
     ELSIF (#tempPostfixNotation[#tempPositionOfPostfix] = #LGCODE_MTH_PRSR_LOGICAL_NOT) THEN
       IF #tempStackOfIntermediateResults[#tempPositionOfIntermediateResult - 1] <> 0 THEN
         #tempStackOfIntermediateResults[#tempPositionOfIntermediateResult - 1] := 0;
       ELSE
         #tempStackOfIntermediateResults[#tempPositionOfIntermediateResult - 1] := 1;
       END_IF;

     ELSIF (#tempPostfixNotation[#tempPositionOfPostfix] = #LGCODE_MTH_PRSR_LOGICAL_NOT_EQUAL) THEN
       IF
         #tempStackOfIntermediateResults[#tempPositionOfIntermediateResult - 2] <>
         #tempStackOfIntermediateResults[#tempPositionOfIntermediateResult - 1]
       THEN
         #tempStackOfIntermediateResults[#tempPositionOfIntermediateResult - 2] := 1;
       ELSE
         #tempStackOfIntermediateResults[#tempPositionOfIntermediateResult - 2] := 0;
       END_IF;
       #tempPositionOfIntermediateResult := #tempPositionOfIntermediateResult - 1;

     ELSIF (#tempPostfixNotation[#tempPositionOfPostfix] = #LGCODE_MTH_PRSR_LOGICAL_EQUAL) THEN
       IF
         #tempStackOfIntermediateResults[#tempPositionOfIntermediateResult - 2] =
         #tempStackOfIntermediateResults[#tempPositionOfIntermediateResult - 1]
       THEN
         #tempStackOfIntermediateResults[#tempPositionOfIntermediateResult - 2] := 1;
       ELSE
         #tempStackOfIntermediateResults[#tempPositionOfIntermediateResult - 2] := 0;
       END_IF;
       #tempPositionOfIntermediateResult := #tempPositionOfIntermediateResult - 1;

     ELSIF (#tempPostfixNotation[#tempPositionOfPostfix] = #LGCODE_MTH_PRSR_LOGICAL_AND) THEN
       IF
         #tempStackOfIntermediateResults[#tempPositionOfIntermediateResult - 2] > 0
         AND
         #tempStackOfIntermediateResults[#tempPositionOfIntermediateResult - 1] > 0
       THEN
         #tempStackOfIntermediateResults[#tempPositionOfIntermediateResult - 2] := 1;
       ELSE
         #tempStackOfIntermediateResults[#tempPositionOfIntermediateResult - 2] := 0;
       END_IF;
       #tempPositionOfIntermediateResult := #tempPositionOfIntermediateResult - 1;

     ELSIF (#tempPostfixNotation[#tempPositionOfPostfix] = #LGCODE_MTH_PRSR_LOGICAL_OR) THEN
       IF
         #tempStackOfIntermediateResults[#tempPositionOfIntermediateResult - 2] > 0
         OR
         #tempStackOfIntermediateResults[#tempPositionOfIntermediateResult - 1] > 0
       THEN
         #tempStackOfIntermediateResults[#tempPositionOfIntermediateResult - 2] := 1;
       ELSE
         #tempStackOfIntermediateResults[#tempPositionOfIntermediateResult - 2] := 0;
       END_IF;
       #tempPositionOfIntermediateResult := #tempPositionOfIntermediateResult - 1;

     END_IF;

     #tempPositionOfPostfix := #tempPositionOfPostfix + 1;

     #LKinLang_CalcMathAndBool.errorID := #LGCODE_MTH_PRSR_NO_ERR;
     #LKinLang_CalcMathAndBool.finalResult := #tempStackOfIntermediateResults[2];

   END_WHILE;

   //--------------------------------------------------------------------
   // End of Block LKinLang_CalcMathAndBool
   //--------------------------------------------------------------------
END_FUNCTION

FUNCTION "LKinLang_CharacterIsLetter" : Bool   // FC35454, SCL
TITLE = LKinLang_CharacterIsLetter
{ S7_Optimized_Access := 'TRUE' }
AUTHOR : tech.team.motioncontrol@siemens.com
FAMILY : LKinLang
VERSION : 1.1
// The FC checks a given character to be a letter
   VAR_INPUT
      character : Byte;   // character to be checked / character to be checked to be a letter
   END_VAR
   // Ret_Val : TRUE: character is letter; FALSE: character is NOT a letter
BEGIN
   //==========================================================================================
   // SIEMENS AG
   // (c)Copyright 2019 All Rights Reserved
   //------------------------------------------------------------------------------------------
   // Library: LKinLang
   // Tested with: S7-1517T-3 PN/DP
   // Engineering: TIA Portal V15
   // Restrictions: ---
   // Requirements: S7-1500T FW 2.5
   // Functionality: LKinLang_CharacterIsLetter
   // The FC checks a given character to be a letter 
   // 
   // Support: tech.team.motioncontrol@siemens.com
   // Note: Parameter comments are only available in language 'English (United States)'
   //------------------------------------------------------------------------------------------
   // Change log table:
   // Version    Date          Expert in charge    Changes applied
   // 01.00.00   28.05.2019    FR                  First created version
   // 01.01.00   09.01.2020    FR                  Added % as letter for interface vars
   //===========================================================================================

   //======================================================================
   // Check if the given characteracter is a LETTER
   //====================================================================== 

                      // A ..................... Z         
   IF ((#character >= 16#41 AND #character <= 16#5A) OR
                    // a ..................... z         
     (#character >= 16#61 AND #character <= 16#7A))
     OR #character = 16#25 //%
   THEN
     #LKinLang_CharacterIsLetter:= TRUE;
   ELSE
     #LKinLang_CharacterIsLetter := FALSE;
   END_IF;
END_FUNCTION

FUNCTION "LKinLang_CharacterIsMerger" : Bool   // FC35455, SCL
TITLE = LKinLang_CharacterIsMerger
{ S7_Optimized_Access := 'TRUE' }
AUTHOR : tech.team.motioncontrol@siemens.com
FAMILY : LKinLang
VERSION : 1.1
// The FC checks a given character to be a merger
   VAR_INPUT
      character : Byte;   // character to be checked
      lastIndexOfMerger : Int;
   END_VAR
   VAR_IN_OUT
      mergers : Array[1.."LKINLANG_NUMBER_OF_MERGERS"] of Byte;
   END_VAR
   VAR_TEMP
      tempCounter : Int;
   END_VAR
   // Ret_Val : TRUE: character is merger; FALSE: character is NOT a merger
BEGIN
   //==========================================================================================
   // SIEMENS AG
   // (c)Copyright 2019 All Rights Reserved
   //------------------------------------------------------------------------------------------
   // Library: LKinLang
   // Tested with: S7-1517T-3 PN/DP
   // Engineering: TIA Portal V15
   // Restrictions: ---
   // Requirements: S7-1500T FW 2.5
   // Functionality: LKinLang_CharacterIsMerger
   // The FC checks a given character to be a merger 
   // 
   // Support: tech.team.motioncontrol@siemens.com
   // Note: Parameter comments are only available in language 'English (United States)'
   //------------------------------------------------------------------------------------------
   // Change log table:
   // Version    Date          Expert in charge    Changes applied
   // 01.00.00   28.05.2019    FR                  First created version
   //===========================================================================================

   //======================================================================
   // Check if the given character is a merger
   //====================================================================== 

   #LKinLang_CharacterIsMerger := false;

   FOR #tempCounter := 1 TO #lastIndexOfMerger DO
     IF #mergers[#tempCounter] = #character THEN
       #LKinLang_CharacterIsMerger := true;
       EXIT;
     END_IF;
   END_FOR;
END_FUNCTION

FUNCTION "LKinLang_CharacterIsNumeric" : Bool   // FC35456, SCL
TITLE = LKinLang_CharacterIsNumeric
{ S7_Optimized_Access := 'TRUE' }
AUTHOR : tech.team.motioncontrol@siemens.com
FAMILY : LKinLang
VERSION : 1.1
// The FC checks a given character to be a numeric
   VAR_INPUT
      character : Char;   // character to be checked
   END_VAR
   // Ret_Val : TRUE: character is numeric; FALSE: character is NOT a numeric
BEGIN
   //==========================================================================================
   // SIEMENS AG
   // (c)Copyright 2019 All Rights Reserved
   //------------------------------------------------------------------------------------------
   // Library: LKinLang
   // Tested with: S7-1517T-3 PN/DP
   // Engineering: TIA Portal V15
   // Restrictions: ---
   // Requirements: S7-1500T FW 2.5
   // Functionality: LKinLang_CharacterIsNumeric
   // The FC checks a given character to be a numeric
   // 
   // Support: tech.team.motioncontrol@siemens.com
   // Note: Parameter comments are only available in language 'English (United States)'
   //------------------------------------------------------------------------------------------
   // Change log table:
   // Version    Date          Expert in charge    Changes applied
   // 01.00.00   28.05.2019    FR                  First created version
   //===========================================================================================

   //======================================================================
   // Check if the given character is a DIGIT or a POINT (used for comma)
   //====================================================================== 

   IF #character = '0'//16#30   // 0
     OR #character = '1'//16#31 // 1
     OR #character = '2'//16#32 // 2
     OR #character = '3'//16#33 // 3
     OR #character = '4'//16#34 // 4
     OR #character = '5'//16#35 // 5
     OR #character = '6'//16#36 // 6
     OR #character = '7'//16#37 // 7 
     OR #character = '8'//16#38 // 8
     OR #character = '9'//16#39 // 9 
     OR #character = '.'//16#2E // .
   THEN
     #LKinLang_CharacterIsNumeric := TRUE;
   ELSE
     #LKinLang_CharacterIsNumeric := FALSE;
   END_IF;
END_FUNCTION

FUNCTION "LKinLang_CheckLimits" : DWord   // FC35457, SCL
TITLE = LKinLang_CheckLimits
{ S7_Optimized_Access := 'TRUE' }
AUTHOR : tech.team.motioncontrol@siemens.com
FAMILY : LKinLang
VERSION : 1.1
// The FC checks a parameter value not to exceed give limits
   VAR_INPUT
      parameterMinVal : LReal;   // lower limit for parameter value
      parameterMaxVal : LReal;   // upper limit for parameter value
   END_VAR
   VAR_IN_OUT
      parameterValue : "LKinLang_typeDiffElementaryDatatypes";   // parameter value which is checked and written
   END_VAR
   VAR CONSTANT
      REAL_MIN : LReal := -3.402823E+38;
      REAL_MAX : LReal := 3.402823E+38;
      DINT_MIN : DInt := -2147483648;
      DINT_MAX : DInt := +2147483647;
      INT_MIN : Int := -32768;
      INT_MAX : Int := 32767;
      ERR_PARAMETER_OVERFLOW : DWord := 16#8000;
      ERR_PARAMETER_OUTSIDE_LIMITS : DWord := 16#8001;
   END_VAR
BEGIN
   //==========================================================================================
   // SIEMENS AG
   // (c)Copyright 2019 All Rights Reserved
   //------------------------------------------------------------------------------------------
   // Library: LKinLang
   // Tested with: S7-1517T-3 PN/DP
   // Engineering: TIA Portal V15
   // Restrictions: ---
   // Requirements: S7-1500T FW 2.5
   // Functionality: LKinLang_CheckLimits
   // The FC checks a parameter value not to exceed give limits
   // 
   // Support: tech.team.motioncontrol@siemens.com
   // Note: Parameter comments are only available in language 'English (United States)'
   //------------------------------------------------------------------------------------------
   // Change log table:
   // Version    Date          Expert in charge    Changes applied
   // 01.00.00   28.05.2019    FR                  First created version
   //===========================================================================================

   // ============================================================
   // Check limits of given parameter
   // ============================================================
   #LKinLang_CheckLimits := 0;

   // Check if parameter value is inside configured limits
   IF #parameterValue.valueLReal >= #parameterMinVal
     AND #parameterValue.valueLReal <= #parameterMaxVal
   THEN
     ; // Value is ok
   ELSE
     ; // Error: Value outside limits  
     #LKinLang_CheckLimits := #ERR_PARAMETER_OUTSIDE_LIMITS;
     RETURN;
   END_IF;

   // Check if parameter value (LReal) fits into smaller data types
   IF #parameterMinVal >= #REAL_MIN
     AND #parameterMaxVal <= #REAL_MAX
   THEN
     // Limits are OK
     IF #parameterValue.valueLReal <= #REAL_MAX
       AND #parameterValue.valueLReal >= #REAL_MIN
     THEN
       #parameterValue.valueReal := LREAL_TO_REAL(#parameterValue.valueLReal);
     ELSE
       // Error
       #LKinLang_CheckLimits := #ERR_PARAMETER_OVERFLOW;
       RETURN;
     END_IF;
   ELSE
     ;// Do nothing: because of the limits this format is not needed
   END_IF;

   IF #parameterMinVal >= #DINT_MIN
     AND #parameterMaxVal <= #DINT_MAX
   THEN
     // Limits are OK
     IF #parameterValue.valueLReal <= #DINT_MAX
       AND #parameterValue.valueLReal >= #DINT_MIN
     THEN
       #parameterValue.valueDint := LREAL_TO_DINT(#parameterValue.valueLReal);
     ELSE
       // Error
       #LKinLang_CheckLimits := #ERR_PARAMETER_OVERFLOW;
       RETURN;
     END_IF;
   ELSE
     ;// Do nothing: because of the limits this format is not needed
   END_IF;

   IF #parameterMinVal >= #INT_MIN
     AND #parameterMaxVal <= #INT_MAX
   THEN
     // Limits are OK
     IF #parameterValue.valueLReal <= #INT_MAX
       AND #parameterValue.valueLReal >= #INT_MIN
     THEN
       #parameterValue.valueInt := LREAL_TO_INT(#parameterValue.valueLReal);
     ELSE
       // Error
       #LKinLang_CheckLimits := #ERR_PARAMETER_OVERFLOW;
       RETURN;
     END_IF;
   ELSE
     ;// Do nothing: because of the limits this format is not needed
   END_IF;
END_FUNCTION

FUNCTION "LKinLang_CheckParameterCondition" : Bool   // FC35458, SCL
TITLE = LKinLang_CheckParameterCondition
{ S7_Optimized_Access := 'TRUE' }
AUTHOR : tech.team.motioncontrol@siemens.com
FAMILY : LKinLang
VERSION : 1.1
// The FC checks for conditions to be fullfilled
   VAR_INPUT
      mode : DInt;   // Selected mode, where the parameters are to be checked (0: In line, 1: In Cmd, 2: In Prg)
      language : Int;   // Selected language
   END_VAR
   VAR_OUTPUT
      errorString : String;   // Generated error message
   END_VAR
   VAR_IN_OUT
      setParameters : Array[1.."LKINLANG_NUMBER_OF_CONDITIONS"] of "LKinLang_typeCondition";   // Array containint all parameters which are set for the selected mode
      conditionsToCheck : Array[1.."LKINLANG_NUMBER_OF_CONDITIONS"] of "LKinLang_typeCondition";   // Array containing all parameters which are to be checked
      parameterDefaults : Variant;   // Parameter defaults to call SelectLangPackage
   END_VAR
   VAR_TEMP
      tempParameterOk : Bool;   // Temporary variable for the return value of this FC
      tempGroupToCheck : DInt;   // Temporary variable for the group which is checked
      tempParameterToCheck : DInt;   // Temporary variable for the parameter number which is checked
      tempConditionCounter : Int;   // Temporary counter in the conditions array
      tempSetCounter : Int;   // Temporary counter in the parameters array
      tempConditionUpperLimit : DInt;   // Temporary variable for upper limit of conditions array
      tempConditionLowerLimit : DInt;   // Temporary variable for lower limit of conditions array
      tempSetUpperLimit : DInt;   // Temporary variable for upper limit of parameters array
      tempSetLowerLimit : DInt;   // Temporary variable for lower limit of parameters array
      tempGroups : Array[1.."LKINLANG_NUMBER_OF_CONDITIONS"] of DInt;   // Temporay array for all groups to be checked
      tempGroupCounter : DInt;   // Temporary variable for last entry in groups array
      tempCounter : Int;   // Temporary counter
      tempParameterDefinition : "LKinLang_typeParameterDefinition";   // Temporary variable for the parameter definition
      tempSep : Array[1.."LKINLANG_NUMBER_OF_SEPARATORS"] of Byte;   // Temporary variable for separators array
      tempMerg : Array[1.."LKINLANG_NUMBER_OF_MERGERS"] of Byte;   // Temporary variable for mergers array
      tempValidCounts : "LKinLang_typePathDataElementCounter";   // Temporary variable for valid counts array
      tempString : "LKinLang_typeVariableDeclaration";
      tempKeyToken : "LKinLang_typeKeyToken";
   END_VAR
   // Ret_Val : Return value of this FC
BEGIN
   //==========================================================================================
   // SIEMENS AG
   // (c)Copyright 2019 All Rights Reserved
   //------------------------------------------------------------------------------------------
   // Library: LKinLang
   // Tested with: S7-1517T-3 PN/DP
   // Engineering: TIA Portal V15
   // Restrictions: ---
   // Requirements: S7-1500T FW 2.5
   // Functionality: LKinLang_CheckParameterCondition
   // This function searches the array "SetParameters" if the parameter number from "ConditionsToCheck" is set.
   // For each group ("conditionsToCheck.Group") there must be at least one parameter number in "SetParameters".
   // 
   // The mode to check is given as an Input:
   // 0: "SetParameters" in the actual line are checked
   // 1: "SetParameters" in the actual command are checked
   // 2: "SetParameters" in the complete program are checked
   // The respective "SetParameters" array must be connected outside
   // 
   // Support: tech.team.motioncontrol@siemens.com
   // Note: Parameter comments are only available in language 'English (United States)'
   //------------------------------------------------------------------------------------------
   // Change log table:
   // Version    Date          Expert in charge    Changes applied
   // 01.00.00   28.05.2019    FR                  First created version
   //===========================================================================================

   // Init variables
   #tempParameterOk := #LKinLang_CheckParameterCondition := FALSE;
   #tempGroupCounter := 0;

   // Get limits of "conditionToCheck" array
   #tempConditionLowerLimit := 1;
   #tempConditionUpperLimit := "LKINLANG_NUMBER_OF_CONDITIONS";

   // Get limits of "setParameters" array
   #tempSetLowerLimit := 1;
   #tempSetUpperLimit := "LKINLANG_NUMBER_OF_CONDITIONS";

   // Iterate over condition array and get all groups which are to be checked
   FOR #tempCounter := #tempConditionLowerLimit TO #tempConditionUpperLimit DO
     // Get group to check
     IF #conditionsToCheck[#tempCounter].Group <> 0 // Group is not 0
       AND #tempGroupToCheck <> #conditionsToCheck[#tempCounter].Group // Group is different from already added group
       AND #conditionsToCheck[#tempCounter].Mode = #mode // Mode is same as selected input
     THEN
       // Increment counter for found groups 
       #tempGroupCounter += 1;
       // Save group number in temp for check in next iteration
       #tempGroupToCheck := #conditionsToCheck[#tempCounter].Group;
       // Save group in array to work with later
       #tempGroups[#tempGroupCounter] := #conditionsToCheck[#tempCounter].Group;
     END_IF;
   END_FOR;

   // Iterate over all found groups ("tempGroups")
   FOR #tempCounter := 1 TO #tempGroupCounter DO
     // Reset Parameter ok
     #tempParameterOk := FALSE;
     // Reset parameter number to check
     #tempParameterToCheck := -1;

     // Search if one group member (parameterNumber) is in "SetParameters" Array 
     FOR #tempConditionCounter := #tempConditionLowerLimit TO #tempConditionUpperLimit DO

       // Search for entries in conditionsToCheck array where ".Group" fits "tempGroups" 
       IF #conditionsToCheck[#tempConditionCounter].Group = #tempGroups[#tempCounter] THEN
         // Group is same --> Get parameter number to check
         #tempParameterToCheck := #conditionsToCheck[#tempConditionCounter].ParameterNumber;
       END_IF;

       // Search in array "SetParameters" if there is an entry which fits the parameterToCheck
       FOR #tempSetCounter := #tempSetLowerLimit TO #tempSetUpperLimit DO
         IF #tempParameterToCheck = #setParameters[#tempSetCounter].ParameterNumber THEN
           // Parameter number was found --> Set parameter ok to True and exit this for Loop
           #tempParameterOk := true;
           EXIT;
         END_IF;
       END_FOR;

       // If one of the group members was found also exit this for loop
       IF #tempParameterOk THEN
         EXIT;
       END_IF;
     END_FOR;

     // If parameter number was not found, generate error message
     IF NOT #tempParameterOk THEN
       // Parameter / Group is missing 
       #errorString := 'Mandatory parameter ';

       FOR #tempConditionCounter := #tempConditionLowerLimit TO #tempConditionUpperLimit DO
         // Get parameter number in conditions to check array, where group fits
         IF #conditionsToCheck[#tempConditionCounter].Group = #tempGroups[#tempCounter] THEN

           // Copy found parameter number
           #tempParameterToCheck := #conditionsToCheck[#tempConditionCounter].ParameterNumber;

           // Get definition of parameter with this number
           "LKinLang_SelectLangPackage"(language := #language,
                                        variableDeclarations=>#tempString,
                                        keyToken=>#tempKeyToken,
                                        parameterDefinition := #tempParameterDefinition,
                                        separators => #tempSep,
                                        mergers => #tempMerg,
                                        validCounts => #tempValidCounts,
                                        parameterNumber := #tempParameterToCheck,
                                        parameterDefaults := #parameterDefaults);


           // Copy the name of the parameter to the error string
           #errorString := CONCAT(IN1 := #errorString, IN2 := #tempParameterDefinition.parameterNameString);

           IF #tempParameterDefinition.parameterNameNumber <> -1 THEN
             // Concat parameterNameNumber and delete sign from DINT_TO_STRING
             #errorString := CONCAT(IN1 := #errorString, IN2 := DELETE(IN := DINT_TO_STRING(#tempParameterDefinition.parameterNameNumber), L := 1, P := 1));
           END_IF;
           // Seperate parameters from the same group with ", "
           #errorString := CONCAT(IN1 := #errorString, IN2 := ', ');
         END_IF;

       END_FOR;
       // Delete last ", "
       #errorString := LEFT(IN := #errorString, L := LEN(#errorString) - 2);
       // Concat last strings
       #errorString := CONCAT(IN1 := #errorString, IN2 := ' is missing');
       // The resulting errorString should look like this
       // "Mandatory parameter G17, G18, G19 is missing" (G17, G18, G19 are for example in the same condition group)
       // 
       // Return from this function
       RETURN;

     ELSE
       // Reset parameter ok for the next group to check
       #tempParameterOk := false;
     END_IF;

   END_FOR;

   // If all groups are ok set parameterOk to true
   // We can assume all parameters were ok because else we would have returned after writing the error string
   #tempParameterOk := true;

   // Write internal temp to output
   #LKinLang_CheckParameterCondition := #tempParameterOk;

   //===========================================================================================
   // End of Block
   //===========================================================================================
END_FUNCTION

FUNCTION "LKinLang_CheckParameterCounter" : Void   // FC35459, SCL
TITLE = LKinLang_CheckParameterCounter
{ S7_Optimized_Access := 'TRUE' }
AUTHOR : tech.team.motioncontrol@siemens.com
FAMILY : LKinLang
VERSION : 1.1
// This function checks how often a parameter was programmed in one line
   VAR_INPUT
      parameterNumber : Int;   // Parameter number for which the counter is checked
      lineNo : UInt;   // Actual line number for error message
      parameterDefinition : "LKinLang_typeParameterDefinition";   // Parameter definition of the parameter number
   END_VAR
   VAR_IN_OUT
      parameterCounter : Array[*] of "LKinLang_typeParameterCounter";   // Parameter counter array
      errorString : String;   // Error message
      error : Bool;   // Error output
   END_VAR
   VAR_TEMP
      tempCounter : Int;   // Temporary counter
      tempUBound : DInt;   // Temporary variable for the upper limit of the parameterCounter array
      tempLBound : DInt;   // Temporary variable for the lower limit of the parameterCounter array
      tempParameterFound : Bool;   // Temporary bit to signalize if the parameter is already in the parameterCounter array
   END_VAR
   // Ret_Val : No return value
BEGIN
   //==========================================================================================
   // SIEMENS AG
   // (c)Copyright 2019 All Rights Reserved
   //------------------------------------------------------------------------------------------
   // Library: LKinLang
   // Tested with: S7-1517T-3 PN/DP
   // Engineering: TIA Portal V15
   // Restrictions: ---
   // Requirements: S7-1500T FW 2.5
   // Functionality: LKinLang_CheckParameterCounter
   // This function checks how often a given parameter was programmed in one line.
   // It increases the counter or throws an error if the limit is exceeded.
   //
   // Support: tech.team.motioncontrol@siemens.com
   // Note: Parameter comments are only available in language 'English (United States)'
   //------------------------------------------------------------------------------------------
   // Change log table:
   // Version    Date          Expert in charge    Changes applied
   // 01.00.00   28.05.2019    FR                  First created version
   //===========================================================================================

   // Initialize variables
   //------------------------------------------------------------------------------------------
   #tempLBound := LOWER_BOUND(ARR := #parameterCounter, DIM := 1);
   #tempUBound := UPPER_BOUND(ARR := #parameterCounter, DIM := 1);
   #tempParameterFound := FALSE;
   //------------------------------------------------------------------------------------------

   // Check if parameter number is already in array
   //------------------------------------------------------------------------------------------
   FOR #tempCounter := #tempLBound TO #tempUBound DO

     // Parameter number is already in array
     IF #parameterCounter[#tempCounter].parameterNumber = #parameterNumber THEN

       // Already in array --> Count up
       #parameterCounter[#tempCounter].counterValue += 1;
       // Set bit to skip creating a new entry
       #tempParameterFound := TRUE;

       // ERROR: Throw error if limit of counter was exceeded
       //------------------------------------------------------------------------------------------
       IF #parameterCounter[#tempCounter].counterValue > #parameterDefinition.validCountPerLine THEN

         // Create error string
         //------------------------------------------------------------------------------------------
         #errorString := CONCAT(IN1 := #errorString, IN2 := 'Programmed ');
         #errorString := CONCAT(IN1 := #errorString, IN2 := #parameterDefinition.parameterNameString);

         // Concat parameterNameNumber if not -1
         // If the parameter does not include a number, e.g. LIN (compared to G2) the parameterNameNumber is -1 by default 
         IF #parameterDefinition.parameterNameNumber <> -1 THEN
           #errorString := CONCAT(IN1 := #errorString, IN2 := DINT_TO_STRING(#parameterDefinition.parameterNameNumber));
         END_IF;
         #errorString := CONCAT(IN1 := #errorString, IN2 := ' too often: Allowed:');
         #errorString := CONCAT(IN1 := #errorString, IN2 := DINT_TO_STRING(#parameterDefinition.validCountPerLine));
         #errorString := CONCAT(IN1 := #errorString, IN2 := ' Programmed:');
         #errorString := CONCAT(IN1 := #errorString, IN2 := INT_TO_STRING(#parameterCounter[#tempCounter].counterValue));
         #errorString := CONCAT(IN1 := #errorString, IN2 := '; Line:');
         #errorString := CONCAT(IN1 := #errorString, IN2 := UINT_TO_STRING(#lineNo));

         // Completed errorString should look like
         // "Programmed G1 too often: Allowed:+1 Programmed: +2; Line:+10 "
         //------------------------------------------------------------------------------------------

         // Set error output to TRUE;
         #error := TRUE;

         // Return from function after errorString is written
         RETURN;
       ELSE
         // Exit for loop if parameter was found and counter was sucessfully increased
         EXIT;
       END_IF;
     ELSE
       ; // Do nothing --> next iteration
     END_IF;
   END_FOR;
   //------------------------------------------------------------------------------------------

   // If parameter was not found, create new entry in parameterCounter array
   //------------------------------------------------------------------------------------------
   IF NOT #tempParameterFound THEN
     // New entry
     // Search empty array index
     FOR #tempCounter := #tempLBound TO #tempUBound DO

       // If CounterValue = 0 then this must be a empty index
       IF #parameterCounter[#tempCounter].counterValue = 0 THEN

         // New entry
         #parameterCounter[#tempCounter].parameterNumber := #parameterNumber;
         // Increment counter
         #parameterCounter[#tempCounter].counterValue += 1;

         // ERROR: Throw error if limit of counter was exceeded
         //------------------------------------------------------------------------------------------
         IF #parameterCounter[#tempCounter].counterValue > #parameterDefinition.validCountPerLine THEN

           // Create error string
           //------------------------------------------------------------------------------------------
           #errorString := CONCAT(IN1 := #errorString, IN2 := 'Programmed ');
           #errorString := CONCAT(IN1 := #errorString, IN2 := #parameterDefinition.parameterNameString);
           // Concat parameterNameNumber if not -1
           // If the parameter does not include a number, e.g. LIN (compared to G2) the parameterNameNumber is -1 by default 
           IF #parameterDefinition.parameterNameNumber <> -1 THEN
             #errorString := CONCAT(IN1 := #errorString, IN2 := DINT_TO_STRING(#parameterDefinition.parameterNameNumber));
           END_IF;
           #errorString := CONCAT(IN1 := #errorString, IN2 := ' too often: Allowed:');
           #errorString := CONCAT(IN1 := #errorString, IN2 := DINT_TO_STRING(#parameterDefinition.validCountPerLine));
           #errorString := CONCAT(IN1 := #errorString, IN2 := ' Programmed:');
           #errorString := CONCAT(IN1 := #errorString, IN2 := INT_TO_STRING(#parameterCounter[#tempCounter].counterValue));
           #errorString := CONCAT(IN1 := #errorString, IN2 := '; Line:');
           #errorString := CONCAT(IN1 := #errorString, IN2 := UINT_TO_STRING(#lineNo));

           // Completed errorString should look like
           // "Programmed G1 too often: Allowed:+1 Programmed: +2; Line:+10 "
           //------------------------------------------------------------------------------------------

           // Set error output to TRUE;
           #error := TRUE;

           // Return from function after errorString is written
           RETURN;
         ELSE
           // Exit for loop if parameter was found and counter was sucessfully increased
           EXIT;
         END_IF;
       ELSE
         ; // Do nothing --> next iteration
       END_IF;
     END_FOR;
     //------------------------------------------------------------------------------------------
   ELSE
     ; // Do nothing --> parameter was found before
   END_IF;

   //===========================================================================================
   // End of Block
   //===========================================================================================
END_FUNCTION

FUNCTION "LKinLang_CheckPathDataCmd" : Word   // FC35460, SCL
TITLE = LKinCtrl_CheckPathDataCmd
{ S7_Optimized_Access := 'TRUE' }
AUTHOR : tech.team.motioncontrol@siemens.com
FAMILY : LKinCtrl
VERSION : 1.1
// The FC checks a PathData command to be configured correctly
   VAR_IN_OUT
      errorString : String;
      pathDataCmd : "LKinCtrl_typePathDataElement_advanced";   // variant for PathData command
   END_VAR
   VAR_TEMP
      tmpError : Bool;   // temporary variable for error bit
      tempFlagCtr : Int;   // temporary counter for flags
   END_VAR
   VAR CONSTANT
      STATUS_NO_ERROR_IN_COMMAND : Word := 16#0000;   // status no error found command
      ERR_PATHDATA_CMDTYPE : Word := 16#80A0;   // error due to wrong cmdType
      ERR_PATHDATA_COORDSYSTEM : Word := 16#80B1;   // error due to wrong coordinate system
      ERR_PATHDATA_ORIENTATIONDIRECTION : Word := 16#8007;   // error due to wrong orientation direction
      ERR_PATHDATA_BUFFERMODE : Word := 16#80B2;   // error due to wrong buffer mode
      ERR_PATHDATA_DYNAMICADAPTION : Word := 16#80B5;   // error due to wrong dynamic adaption
      ERR_PATHDATA_CIRCMODE : Word := 16#80B6;   // error due to wrong circle mode
      ERR_PATHDATA_PATHCHOICE : Word := 16#80B9;   // error due to wrong path choice
      ERR_PATHDATA_CIRCLEPLANE : Word := 16#80BA;   // error due to wrong circle plane
      ERR_PATHDATA_RADIUS : Word := 16#80BB;   // error due to wrong radius
      ERR_PATHDATA_ARC : Word := 16#80BC;   // error due to wrong arc
      ERR_PATHDATA_SETFLAGS_FLAG : Word := 16#80D1;   // error due to wrong flag definition
      ERR_PATHDATA_SETFLAGS_FLAGMODE : Word := 16#80D2;   // error due to wrong flag mode definition / errot due to wrong flag mode definition
      ERR_PATHDATA_OFFSET_PARA_NO : Word := 16#80A1;   // error due to wrong offset parameter set number / errot due to wrong offset parameter set number
      ERR_PATHDATA_OFFSET_MAINPATHPLANE : Word := 16#80A2;   // error due to wrong main path plane
      MINVAL_LREAL : LReal := -1.7976931348623157E+308;
      MINVAL_DINT : DInt := -2_147_483_648;
      MINVAL_INT : Int := -32_768;
   END_VAR
BEGIN
   //==========================================================================================
   // SIEMENS AG
   // (c)Copyright 2019 All Rights Reserved
   //------------------------------------------------------------------------------------------
   // Library: LKinLang
   // Tested with: S7-1517T-3 PN/DP
   // Engineering: TIA Portal V15
   // Restrictions: ---
   // Requirements: S7-1500T FW 2.5
   // Functionality: LKinLang_CheckPathDataCmd
   // The FC checks a PathData command to be configured correctly
   // 
   // Support: tech.team.motioncontrol@siemens.com
   // Note: Parameter comments are only available in language 'English (United States)'
   //------------------------------------------------------------------------------------------
   // Change log table:
   // Version    Date          Expert in charge    Changes applied
   // 01.00.00   28.05.2019    FR                  First created version
   // 01.00.01   26.11.2019    FR                  Added flagOnly cmd to CmdType check; added value Flags
   // 01.00.02   12.02.2020    FR                  Use correct constant for valueFlags
   // 01.00.03   10.12.2020    FR                  Check for cmdType=-1 
   //===========================================================================================

   // FC initialization
   //====================================================================================================================================
   #tmpError := FALSE;
   #LKinLang_CheckPathDataCmd := #STATUS_NO_ERROR_IN_COMMAND;

   // PathData command 
   //====================================================================================================================================
   //PathData - command - cmdType
   // Check for cmdType = -1 
   // This FC is only called to check valid motion commands
   // => -1 is not allowed
   // => End of PathData is written in other step
   IF #pathDataCmd.cmdType = -1 THEN
       #tmpError := TRUE;
       #LKinLang_CheckPathDataCmd := #ERR_PATHDATA_CMDTYPE;
       #errorString := CONCAT(IN1 := #errorString, IN2 := 'Error: Missing motion command');
       RETURN;
   END_IF;


   // check for wrong PathData parameter cmdType
   IF (#pathDataCmd.cmdType < "LKINCTRL_CMD_FLAG_ONLY"                      // lower limit MC cmdTypes
     OR #pathDataCmd.cmdType > "LKINCTRL_MC_MOVECIRCULARREL")               // upper limit MC cmdTypes
     AND #pathDataCmd.cmdType <> "LKINCTRL_CMD_WAIT_TIME"                   // exact cmdType constant for wait time
     AND #pathDataCmd.cmdType <> "LKINCTRL_CONFIG_START_OFFSET_COMP_LEFT"   // exact cmdType constant for activation offset compensation left
     AND #pathDataCmd.cmdType <> "LKINCTRL_CONFIG_START_OFFSET_COMP_RIGHT"  // exact cmdType constant for activation offset compensation right
     AND #pathDataCmd.cmdType <> "LKINCTRL_CONFIG_END_OFFSET_COMP"          // exact cmdType constant for deactivation offset compensation
   THEN
     #tmpError := TRUE;
     #LKinLang_CheckPathDataCmd := #ERR_PATHDATA_CMDTYPE;
     #errorString := CONCAT(IN1 := #errorString, IN2 := 'Error: cmdType = ');
     #errorString := CONCAT(IN1 := #errorString, IN2 := INT_TO_STRING(#pathDataCmd.cmdType));
     #errorString := CONCAT(IN1 := #errorString, IN2 := ' not allowed');
     RETURN;
   END_IF;


   //PathData - command - cmdCoordinates - coordSystem
   // check for wrong parameter PathData coordSystem
   IF #pathDataCmd.cmdCoordinates.coordSystem < 0
     AND #pathDataCmd.cmdCoordinates.coordSystem > 3
   THEN
     #tmpError := TRUE;
     #LKinLang_CheckPathDataCmd := #ERR_PATHDATA_COORDSYSTEM;
     #errorString := CONCAT(IN1 := #errorString, IN2 := 'Error: Coordinate system = ');
     #errorString := CONCAT(IN1 := #errorString, IN2 := DINT_TO_STRING(#pathDataCmd.cmdCoordinates.coordSystem));
     #errorString := CONCAT(IN1 := #errorString, IN2 := ' not allowed');
     RETURN;
   END_IF;

   //PathData - command - cmdParameters - orientationDirection
   // check for wrong parameter PathData orientationDirection
   IF #pathDataCmd.cmdParameters.orientationDirection < 1
     OR #pathDataCmd.cmdParameters.orientationDirection > 3
   THEN
     #tmpError := TRUE;
     #LKinLang_CheckPathDataCmd := #ERR_PATHDATA_ORIENTATIONDIRECTION;
     #errorString := CONCAT(IN1 := #errorString, IN2 := 'Error: Orientation direction = ');
     #errorString := CONCAT(IN1 := #errorString, IN2 := DINT_TO_STRING(#pathDataCmd.cmdParameters.orientationDirection));
     #errorString := CONCAT(IN1 := #errorString, IN2 := ' not allowed');
     RETURN;
   END_IF;

   //PathData - command - cmdParameters - bufferMode
   // check for wrong parameter PathData bufferMode
   IF #pathDataCmd.cmdParameters.bufferMode <> 1
     AND #pathDataCmd.cmdParameters.bufferMode <> 2
     AND #pathDataCmd.cmdParameters.bufferMode <> 5
   THEN
     #tmpError := TRUE;
     #LKinLang_CheckPathDataCmd := #ERR_PATHDATA_BUFFERMODE;
     #errorString := CONCAT(IN1 := #errorString, IN2 := 'Error: Buffer mode = ');
     #errorString := CONCAT(IN1 := #errorString, IN2 := DINT_TO_STRING(#pathDataCmd.cmdParameters.bufferMode));
     #errorString := CONCAT(IN1 := #errorString, IN2 := ' not allowed');
     RETURN;
   END_IF;

   //PathData - command - cmdParameters - dynamicAdaption
   // check for wrong parameter PathData dynamicAdaption
   IF #pathDataCmd.cmdParameters.dynamicAdaption > 2
   THEN
     #tmpError := TRUE;
     #LKinLang_CheckPathDataCmd := #ERR_PATHDATA_DYNAMICADAPTION;
     #errorString := CONCAT(IN1 := #errorString, IN2 := 'Error: Dynamic adaption = ');
     #errorString := CONCAT(IN1 := #errorString, IN2 := DINT_TO_STRING(#pathDataCmd.cmdParameters.dynamicAdaption));
     #errorString := CONCAT(IN1 := #errorString, IN2 := ' not allowed');
     RETURN;
   END_IF;

   //PathData - command - circleParameter
   //====================================================================================================================================
   //PathData - command - circleParameter - circMode
   // check for wrong parameter PathData circMode
   IF #pathDataCmd.cmdParameters.circleParameters.circMode < 0
     OR #pathDataCmd.cmdParameters.circleParameters.circMode > 3
   THEN
     #tmpError := TRUE;
     #LKinLang_CheckPathDataCmd := #ERR_PATHDATA_CIRCMODE;
     #errorString := CONCAT(IN1 := #errorString, IN2 := 'Error: Circle mode = ');
     #errorString := CONCAT(IN1 := #errorString, IN2 := DINT_TO_STRING(#pathDataCmd.cmdParameters.circleParameters.circMode));
     #errorString := CONCAT(IN1 := #errorString, IN2 := ' not allowed');
     RETURN;
   END_IF;

   //PathData - command - circleParameter - pathChoice
   // check for wrong parameter PathData pathChoice
   IF #pathDataCmd.cmdParameters.circleParameters.pathChoice < 0
     OR #pathDataCmd.cmdParameters.circleParameters.pathChoice > 3
   THEN
     #tmpError := TRUE;
     #LKinLang_CheckPathDataCmd := #ERR_PATHDATA_PATHCHOICE;
     #errorString := CONCAT(IN1 := #errorString, IN2 := 'Error: Path choice = ');
     #errorString := CONCAT(IN1 := #errorString, IN2 := DINT_TO_STRING(#pathDataCmd.cmdParameters.circleParameters.pathChoice));
     #errorString := CONCAT(IN1 := #errorString, IN2 := ' not allowed');
     RETURN;
   END_IF;

   //PathData - command - circleParameter - circlePlane
   // check for wrong parameter PathData circlePlane
   IF #pathDataCmd.cmdParameters.circleParameters.circlePlane < 0
     OR #pathDataCmd.cmdParameters.circleParameters.circlePlane > 2
   THEN
     #tmpError := TRUE;
     #LKinLang_CheckPathDataCmd := #ERR_PATHDATA_CIRCLEPLANE;
     #errorString := CONCAT(IN1 := #errorString, IN2 := 'Error: Circle plane = ');
     #errorString := CONCAT(IN1 := #errorString, IN2 := DINT_TO_STRING(#pathDataCmd.cmdParameters.circleParameters.circlePlane));
     #errorString := CONCAT(IN1 := #errorString, IN2 := ' not allowed');
     RETURN;
   END_IF;

   //PathData - command - circleParameter - radius
   // check for wrong parameter PathData radius
   IF #pathDataCmd.cmdParameters.circleParameters.radius < 0.0
   THEN
     #tmpError := TRUE;
     #LKinLang_CheckPathDataCmd := #ERR_PATHDATA_RADIUS;
     #errorString := CONCAT(IN1 := #errorString, IN2 := 'Error: Circle radius = ');
     #errorString := CONCAT(IN1 := #errorString, IN2 := LREAL_TO_STRING(#pathDataCmd.cmdParameters.circleParameters.radius));
     #errorString := CONCAT(IN1 := #errorString, IN2 := ' not allowed');
     RETURN;
   END_IF;

   //PathData - command - circleParameter - arc
   // check for wrong parameter PathData arc
   IF #pathDataCmd.cmdParameters.circleParameters.arc < 0.0
   THEN
     #tmpError := TRUE;
     #LKinLang_CheckPathDataCmd := #ERR_PATHDATA_ARC;
     #errorString := CONCAT(IN1 := #errorString, IN2 := 'Error: Circle arc = ');
     #errorString := CONCAT(IN1 := #errorString, IN2 := LREAL_TO_STRING(#pathDataCmd.cmdParameters.circleParameters.arc));
     #errorString := CONCAT(IN1 := #errorString, IN2 := ' not allowed');
     RETURN;
   END_IF;

   //PathData - command - offsetParameters - offSetParaNo
   // check for wrong parameter offSetParaNo
   IF (#pathDataCmd.cmdType = "LKINCTRL_CONFIG_START_OFFSET_COMP_LEFT"
     OR #pathDataCmd.cmdType = "LKINCTRL_CONFIG_START_OFFSET_COMP_RIGHT")
     AND (#pathDataCmd.cmdParameters.offsetParameters.offsetParaNo < 1
     OR #pathDataCmd.cmdParameters.offsetParameters.offsetParaNo > "LKINCTRL_NO_OF_OFFSETS")
   THEN
     #tmpError := TRUE;
     #LKinLang_CheckPathDataCmd := #ERR_PATHDATA_OFFSET_PARA_NO;
     #errorString := CONCAT(IN1 := #errorString, IN2 := 'Error: Offset parameter number = ');
     #errorString := CONCAT(IN1 := #errorString, IN2 := DINT_TO_STRING(#pathDataCmd.cmdParameters.offsetParameters.offsetParaNo));
     #errorString := CONCAT(IN1 := #errorString, IN2 := ' not allowed');
     RETURN;
   END_IF;

   //PathData - command - offsetParameters - main
   // check for wrong parameter PathData circlePlane
   IF (#pathDataCmd.cmdType = "LKINCTRL_CONFIG_START_OFFSET_COMP_LEFT"
     OR #pathDataCmd.cmdType = "LKINCTRL_CONFIG_START_OFFSET_COMP_RIGHT")
     AND (#pathDataCmd.cmdParameters.offsetParameters.mainPathPlane < 0
     OR #pathDataCmd.cmdParameters.offsetParameters.mainPathPlane > 2)
   THEN
     #tmpError := TRUE;
     #LKinLang_CheckPathDataCmd := #ERR_PATHDATA_OFFSET_MAINPATHPLANE;
     #errorString := CONCAT(IN1 := #errorString, IN2 := 'Error: Offset main path plane = ');
     #errorString := CONCAT(IN1 := #errorString, IN2 := DINT_TO_STRING(#pathDataCmd.cmdParameters.offsetParameters.mainPathPlane));
     #errorString := CONCAT(IN1 := #errorString, IN2 := ' not allowed');
     RETURN;
   END_IF;

   //PathData - command - setFlags
   //====================================================================================================================================
   FOR #tempFlagCtr := 1 TO "LKINCTRL_NO_OF_CMD_SETFLAGS" DO
     // check flag to be in range of flags InOut array at LKinCtrl_MC_MovePath
     IF #pathDataCmd.setFlags[#tempFlagCtr].flag < -1
       OR #pathDataCmd.setFlags[#tempFlagCtr].flag > "LKINCTRL_NO_OF_LAST_SETFLAG"
     THEN
       #tmpError := TRUE;
       #LKinLang_CheckPathDataCmd := #ERR_PATHDATA_SETFLAGS_FLAG;
       #errorString := CONCAT(IN1 := #errorString, IN2 := 'Error: Flag index = ');
       #errorString := CONCAT(IN1 := #errorString, IN2 := DINT_TO_STRING(#pathDataCmd.setFlags[#tempFlagCtr].flag));
       #errorString := CONCAT(IN1 := #errorString, IN2 := ' not allowed');
       EXIT;
       RETURN;
     END_IF;

     // check flagMode to be valid
     IF #pathDataCmd.setFlags[#tempFlagCtr].flagMode <> 0
       AND #pathDataCmd.setFlags[#tempFlagCtr].flagMode <> 1
       AND #pathDataCmd.setFlags[#tempFlagCtr].flagMode <> 2
       AND #pathDataCmd.setFlags[#tempFlagCtr].flagMode <> 3
       AND #pathDataCmd.setFlags[#tempFlagCtr].flagMode <> 5
       AND #pathDataCmd.setFlags[#tempFlagCtr].flagMode <> 10
       AND #pathDataCmd.setFlags[#tempFlagCtr].flagMode <> 11
       AND #pathDataCmd.setFlags[#tempFlagCtr].flagMode <> 13
       AND #pathDataCmd.setFlags[#tempFlagCtr].flagMode <> 15
     THEN
       #tmpError := TRUE;
       #LKinLang_CheckPathDataCmd := #ERR_PATHDATA_SETFLAGS_FLAGMODE;
       #errorString := CONCAT(IN1 := #errorString, IN2 := 'Error: Flag mode = ');
       #errorString := CONCAT(IN1 := #errorString, IN2 := DINT_TO_STRING(#pathDataCmd.setFlags[#tempFlagCtr].flagMode));
       #errorString := CONCAT(IN1 := #errorString, IN2 := ' not allowed');
       EXIT;
       RETURN;
     END_IF;
   END_FOR;

   //PathData - command - valueFlags
   //====================================================================================================================================
   FOR #tempFlagCtr := 1 TO "LKINCTRL_NO_OF_CMD_VALUEFLAGS" DO
     // check flag to be in range of flags InOut array at LKinCtrl_MC_MovePath
     IF #pathDataCmd.valueFlags[#tempFlagCtr].flag < -1
       OR #pathDataCmd.valueFlags[#tempFlagCtr].flag > "LKINCTRL_NO_OF_LAST_VALUEFLAG"
     THEN
       #tmpError := TRUE;
       #LKinLang_CheckPathDataCmd := #ERR_PATHDATA_SETFLAGS_FLAG;
       #errorString := CONCAT(IN1 := #errorString, IN2 := 'Error: Flag index = ');
       #errorString := CONCAT(IN1 := #errorString, IN2 := DINT_TO_STRING(#pathDataCmd.valueFlags[#tempFlagCtr].flag));
       #errorString := CONCAT(IN1 := #errorString, IN2 := ' not allowed');
       EXIT;
       RETURN;
     END_IF;

     // check flagMode to be valid
     IF #pathDataCmd.valueFlags[#tempFlagCtr].flagMode <> 0
       AND #pathDataCmd.valueFlags[#tempFlagCtr].flagMode <> 1
       AND #pathDataCmd.valueFlags[#tempFlagCtr].flagMode <> 2
       AND #pathDataCmd.valueFlags[#tempFlagCtr].flagMode <> 3
       AND #pathDataCmd.valueFlags[#tempFlagCtr].flagMode <> 5
       AND #pathDataCmd.valueFlags[#tempFlagCtr].flagMode <> 10
       AND #pathDataCmd.valueFlags[#tempFlagCtr].flagMode <> 11
       AND #pathDataCmd.valueFlags[#tempFlagCtr].flagMode <> 13
       AND #pathDataCmd.valueFlags[#tempFlagCtr].flagMode <> 15
     THEN
       #tmpError := TRUE;
       #LKinLang_CheckPathDataCmd := #ERR_PATHDATA_SETFLAGS_FLAGMODE;
       #errorString := CONCAT(IN1 := #errorString, IN2 := 'Error: Flag mode = ');
       #errorString := CONCAT(IN1 := #errorString, IN2 := DINT_TO_STRING(#pathDataCmd.valueFlags[#tempFlagCtr].flagMode));
       #errorString := CONCAT(IN1 := #errorString, IN2 := ' not allowed');
       EXIT;
       RETURN;
     END_IF;
   END_FOR;
END_FUNCTION

FUNCTION "LKinLang_CheckProperty" : Bool   // FC35461, SCL
TITLE = LKinLang_CheckProperty
{ S7_Optimized_Access := 'TRUE' }
AUTHOR : tech.team.motioncontrol@siemens.com
FAMILY : LKinLang
VERSION : 1.1
// The FC checks if the given property is set
   VAR_INPUT
      properties : DWord;   // given properties
      propertyToCheck : DWord;   // property to be checked for given properties
   END_VAR
   // Ret_Val : TRUE: property is set; FALSE: property is NOT set
BEGIN
   //==========================================================================================
   // SIEMENS AG
   // (c)Copyright 2019 All Rights Reserved
   //------------------------------------------------------------------------------------------
   // Library: LKinLang
   // Tested with: S7-1517T-3 PN/DP
   // Engineering: TIA Portal V15
   // Restrictions: ---
   // Requirements: S7-1500T FW 2.5
   // Functionality: LKinLang_CheckProperty
   // The FC checks if the given property is set
   // 
   // Support: tech.team.motioncontrol@siemens.com
   // Note: Parameter comments are only available in language 'English (United States)'
   //------------------------------------------------------------------------------------------
   // Change log table:
   // Version    Date          Expert in charge    Changes applied
   // 01.00.00   28.05.2019    FR                  First created version
   //===========================================================================================

